       #STC_PH_xInitializeCard := TRUE;
       #STC_ST_xCardInitialized := FALSE;
   END_IF;
   #_w1 := #STC_ST_xRequestCardInitialization AND NOT #STC_ST_xPhaseInProgress AND NOT #STC_ST_xStoppingFaults AND NOT #INP_tHSCCount.ldStsSlot0;
   IF #_w1 THEN
       #STC_ST_xRequestCardInitialization := FALSE;
       #STC_AUX_tOutHSC.loadValue0 := 0;
   END_IF;
END_REGION

REGION Network 17: End initialize counter card
   RUNG wire#powerrail
      Contact( #STC_PH_xInitializeCard )
      wire#w1
      Contact( #STC_ST_xStoppingFaults )
      wire#w2
      R_Coil( #STC_PH_xInitializeCard )
   END_RUNG
   RUNG wire#w1
      Contact( #INP_tHSCCount.ldStsSlot0 )
   END_RUNG wire#w2
   RUNG wire#w2
      Coil( #STC_PH_xEndInitializeCard )
   END_RUNG
   // the same network as SCL:
   #_w1 := #STC_PH_xInitializeCard AND (#STC_ST_xStoppingFaults OR #INP_tHSCCount.ldStsSlot0);
   IF #_w1 THEN #STC_PH_xInitializeCard := FALSE; END_IF;
   #STC_PH_xEndInitializeCard := #_w1;
END_REGION

REGION Network 18: Set card initialized
   RUNG wire#powerrail
      Contact( #STC_PH_xEndInitializeCard )
      Contact( #INP_tHSCCount.ldStsSlot0 )
      I_Contact( #STC_ST_xStoppingFaults )
      wire#w1
      S_Coil( #STC_ST_xCardInitialized )
   END_RUNG
   RUNG wire#w1
      Coil( #TMP_xInitializeData )
   END_RUNG
   // the same network as SCL:
   #_w1 := #STC_PH_xEndInitializeCard AND #INP_tHSCCount.ldStsSlot0 AND NOT #STC_ST_xStoppingFaults;
   IF #_w1 THEN #STC_ST_xCardInitialized := TRUE; END_IF;
   #TMP_xInitializeData := #_w1;
END_REGION

REGION Network 19 (SCL): Initialize structure after initialization
   IF #TMP_xInitializeData THEN

       #INO_tEncoder.dActualEncoderCounter_cmm := 0;
       #INO_tEncoder.dLastMeterValue_cmm := 0;
       #INO_tEncoder.dNextMeterValue_cmm := #CONST_DMETERINC_CMM;
       #INO_tEncoder.rActSpeedValue_cmm_ms := 0.0;
       #STC_AUX_dLastCounterValue_cmm := 0;

       FOR #TMP_dIndex := 0 TO "DMAXXHEADS_IND" DO
           #INO_tEncoder.rgxMetersForXcuts[#TMP_dIndex] := FALSE;
       END_FOR;

       FOR #TMP_dIndex := 0 TO "DMAXYCUTBRIDGE_IND" DO
           #INO_tEncoder.rgxMetersForYCuts[#TMP_dIndex] := FALSE;
       END_FOR;

       #INO_tEncoder.xMeterForMarkers := FALSE;
       #INO_tEncoder.xMeterForScanner := FALSE;

       #STC_AUX_dLastMeterValue_cmm := 0;
       #STC_AUX_dNextMeterValue_cmm := #CONST_DMETERINC_CMM;
       #STC_AUX_lrTimingCounter_s := 0;
       #STC_AUX_lrTimingCounterFast_s := 0;
       #STC_AUX_dMeterValueSent_cmm := 0;

   END_IF;
END_REGION

REGION Network 20: ####_METER_THRESHOLD_####
END_REGION

REGION Network 21: Update new meter
   RUNG wire#powerrail
      Contact( #STC_ST_xCardInitialized )
      I_Contact( #STC_ST_xRequestCardInitialization )
      I_Contact( #STC_ST_xPhaseInProgress )
      I_Contact( #STC_ST_xStoppingFaults )
      I_Contact( #INP_tHSCCount.ldStsSlot0 )
      { S7_Templates := "SrcType := DInt" } NE_Contact(in1 := #STC_AUX_dNextMeterValue_cmm, in2 := #STC_AUX_dMeterValueSent_cmm)
      wire#w1
      S_Coil( #STC_PH_xUpdateNewMeter )
   END_RUNG
   RUNG wire#w1
      Move(in := #STC_AUX_dNextMeterValue_cmm, out1 => #STC_AUX_tOutHSC.loadValue0)
   END_RUNG
   // the same network as SCL:
   IF #STC_ST_xCardInitialized AND NOT #STC_ST_xRequestCardInitialization AND NOT #STC_ST_xPhaseInProgress AND NOT #STC_ST_xStoppingFaults AND NOT #INP_tHSCCount.ldStsSlot0 AND (#STC_AUX_dNextMeterValue_cmm <> #STC_AUX_dMeterValueSent_cmm) THEN
       #STC_PH_xUpdateNewMeter := TRUE;
       #STC_AUX_tOutHSC.loadValue0 := #STC_AUX_dNextMeterValue_cmm;
   END_IF;
END_REGION

REGION Network 22: End update new meter
   RUNG wire#powerrail
      Contact( #STC_PH_xUpdateNewMeter )
      wire#w1
      Contact( #INP_tHSCCount.ldStsSlot0 )
      wire#w2
      R_Coil( #STC_PH_xUpdateNewMeter )
   END_RUNG
   RUNG wire#w1
      Contact( #IN_xSimulationActive )
   END_RUNG wire#w2
   RUNG wire#w1
      Contact( #STC_ST_xStoppingFaults )
   END_RUNG wire#w2
   RUNG wire#w2
      Coil( #STC_PH_xEndUpdateNewMeter )
   END_RUNG
   // the same network as SCL:
   #_w1 := #STC_PH_xUpdateNewMeter AND (#INP_tHSCCount.ldStsSlot0 OR #IN_xSimulationActive OR #STC_ST_xStoppingFaults);
   IF #_w1 THEN #STC_PH_xUpdateNewMeter := FALSE; END_IF;
   #STC_PH_xEndUpdateNewMeter := #_w1;
END_REGION

REGION Network 23: Set meter correctly written
   RUNG wire#powerrail
      Contact( #STC_PH_xEndUpdateNewMeter )
      wire#w1
      Contact( #INP_tHSCCount.ldStsSlot0 )
      wire#w2
      Move(in := #STC_AUX_dNextMeterValue_cmm, out1 => #STC_AUX_dMeterValueSent_cmm)
   END_RUNG
   RUNG wire#w1
      Contact( #IN_xSimulationActive )
   END_RUNG wire#w2
   // the same network as SCL:
   IF #STC_PH_xEndUpdateNewMeter AND (#INP_tHSCCount.ldStsSlot0 OR #IN_xSimulationActive) THEN
       #STC_AUX_dMeterValueSent_cmm := #STC_AUX_dNextMeterValue_cmm;
   END_IF;
END_REGION

REGION Network 24: ####_NEW METER ARRIVED_####
END_REGION

REGION Network 25: Check if new meter arrived
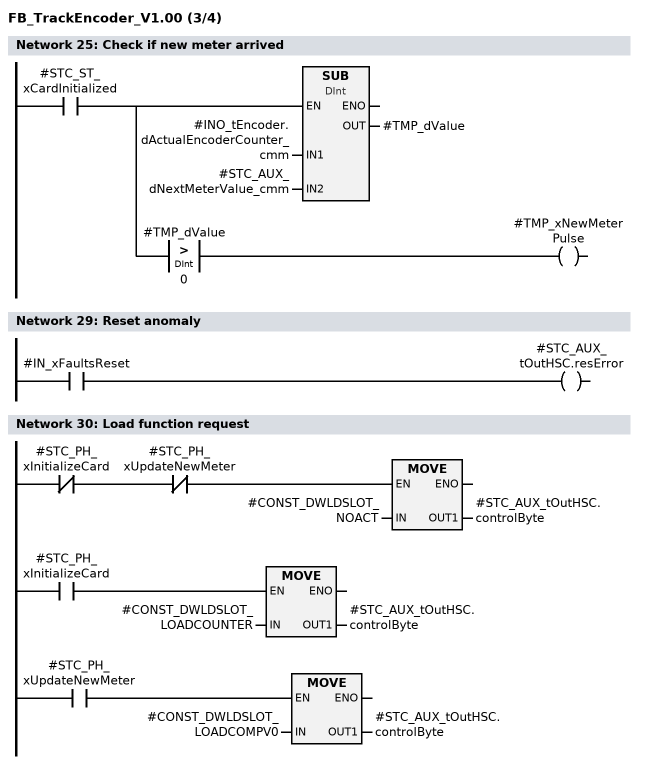
   RUNG wire#powerrail
      Contact( #STC_ST_xCardInitialized )
      wire#w1
      { S7_Templates := "SrcType := DInt" } Sub(in1 := #INO_tEncoder.dActualEncoderCounter_cmm, in2 := #STC_AUX_dNextMeterValue_cmm, out => #TMP_dValue)
   END_RUNG
   RUNG wire#w1
      { S7_Templates := "SrcType := DInt" } GT_Contact(in1 := #TMP_dValue, in2 := 0)
      Coil( #TMP_xNewMeterPulse )
   END_RUNG
   // the same network as SCL:
   IF #STC_ST_xCardInitialized THEN
       #TMP_dValue := #INO_tEncoder.dActualEncoderCounter_cmm - #STC_AUX_dNextMeterValue_cmm;
   END_IF;
   #TMP_xNewMeterPulse := #STC_ST_xCardInitialized AND (#TMP_dValue > 0);
END_REGION

REGION Network 26 (SCL): New meter pulse
   IF #TMP_xNewMeterPulse THEN

       #STC_AUX_dLastMeterValue_cmm := #STC_AUX_dNextMeterValue_cmm;
       #STC_AUX_dNextMeterValue_cmm += #CONST_DMETERINC_CMM;

       #INO_tEncoder.dLastMeterValue_cmm := #STC_AUX_dLastMeterValue_cmm; 
       #INO_tEncoder.dNextMeterValue_cmm := #STC_AUX_dNextMeterValue_cmm; 

       FOR #TMP_dIndex := 0 TO "DMAXXHEADS_IND" DO
           #INO_tEncoder.rgxMetersForXcuts[#TMP_dIndex] := TRUE;
       END_FOR;

       FOR #TMP_dIndex := 0 TO "DMAXYCUTBRIDGE_IND" DO
           #INO_tEncoder.rgxMetersForYCuts[#TMP_dIndex] := TRUE;
       END_FOR;

       #INO_tEncoder.xMeterForMarkers := TRUE;
       #INO_tEncoder.xMeterForScanner := TRUE;


   END_IF;
END_REGION

REGION Network 27 (SCL): Calculate speed
   #STC_AUX_lrTimingCounter_s += #STC_AUX_lrElapsedTime_s;
   #STC_AUX_lrTimingCounterFast_s += #STC_AUX_lrElapsedTime_s;

   IF #STC_AUX_lrTimingCounter_s >= #CONST_LRUPDATESPEED_S THEN

       #TMP_dElapsedPulses_cmm := #INO_tEncoder.dActualEncoderCounter_cmm - #STC_AUX_dLastCounterValue_cmm;

       #INO_tEncoder.rActSpeedValue_cmm_ms := DINT_TO_REAL(#TMP_dElapsedPulses_cmm) / (LREAL_TO_REAL(#STC_AUX_lrTimingCounter_s) * 1000.0);
       #INO_tEncoder.dActSpeedValue_mm_min := REAL_TO_DINT(#INO_tEncoder.rActSpeedValue_cmm_ms * 600.0);    

       #STC_AUX_dLastCounterValue_cmm := #INO_tEncoder.dActualEncoderCounter_cmm;
       #STC_AUX_lrTimingCounter_s := 0;

   END_IF;

   IF #STC_AUX_lrTimingCounterFast_s >= #CONST_LRUPDATESPEEDFAST_S THEN

       #TMP_dElapsedPulses_cmm := #INO_tEncoder.dActualEncoderCounter_cmm - #STC_AUX_dLastCounterValueFast_cmm;

       #INO_tEncoder.rActSpeedValueFast_cmm_ms := DINT_TO_REAL(#TMP_dElapsedPulses_cmm) / (LREAL_TO_REAL(#STC_AUX_lrTimingCounterFast_s) * 1000.0);
       #INO_tEncoder.dActSpeedValueFast_mm_min := REAL_TO_DINT(#INO_tEncoder.rActSpeedValueFast_cmm_ms * 600.0);    

       #STC_AUX_dLastCounterValueFast_cmm := #INO_tEncoder.dActualEncoderCounter_cmm;
       #STC_AUX_lrTimingCounterFast_s := 0;

   END_IF;
END_REGION

REGION Network 28: ####_OUTPUT_####
END_REGION

REGION Network 29: Reset anomaly
   RUNG wire#powerrail
      Contact( #IN_xFaultsReset )
      Coil( #STC_AUX_tOutHSC.resError )
   END_RUNG
   // the same network as SCL:
   #STC_AUX_tOutHSC.resError := #IN_xFaultsReset;
END_REGION

REGION Network 30: Load function request
   RUNG wire#powerrail
      I_Contact( #STC_PH_xInitializeCard )
      I_Contact( #STC_PH_xUpdateNewMeter )
      Move(in := #CONST_DWLDSLOT_NOACT, out1 => #STC_AUX_tOutHSC.controlByte)
   END_RUNG
   RUNG wire#powerrail
      Contact( #STC_PH_xInitializeCard )
      Move(in := #CONST_DWLDSLOT_LOADCOUNTER, out1 => #STC_AUX_tOutHSC.controlByte)
   END_RUNG
   RUNG wire#powerrail
      Contact( #STC_PH_xUpdateNewMeter )
      Move(in := #CONST_DWLDSLOT_LOADCOMPV0, out1 => #STC_AUX_tOutHSC.controlByte)
   END_RUNG
   // the same network as SCL:
   IF NOT #STC_PH_xInitializeCard AND NOT #STC_PH_xUpdateNewMeter THEN
       #STC_AUX_tOutHSC.controlByte := #CONST_DWLDSLOT_NOACT;
   END_IF;
   IF #STC_PH_xInitializeCard THEN #STC_AUX_tOutHSC.controlByte := #CONST_DWLDSLOT_LOADCOUNTER; END_IF;
   IF #STC_PH_xUpdateNewMeter THEN #STC_AUX_tOutHSC.controlByte := #CONST_DWLDSLOT_LOADCOMPV0; END_IF;
END_REGION

REGION Network 31: Fixed command
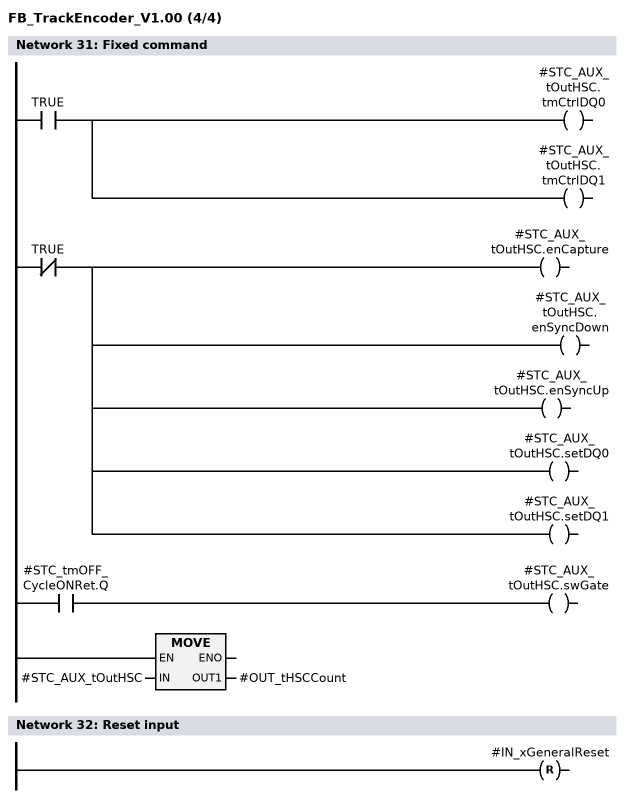
   RUNG wire#powerrail
      Contact( TRUE )
      wire#w1
      Coil( #STC_AUX_tOutHSC.tmCtrlDQ0 )
   END_RUNG
   RUNG wire#w1
      Coil( #STC_AUX_tOutHSC.tmCtrlDQ1 )
   END_RUNG
   RUNG wire#powerrail
      I_Contact( TRUE )
      wire#w2
      Coil( #STC_AUX_tOutHSC.enCapture )
   END_RUNG
   RUNG wire#w2
      Coil( #STC_AUX_tOutHSC.enSyncDown )
   END_RUNG
   RUNG wire#w2
      Coil( #STC_AUX_tOutHSC.enSyncUp )
   END_RUNG
   RUNG wire#w2
      Coil( #STC_AUX_tOutHSC.setDQ0 )
   END_RUNG
   RUNG wire#w2
      Coil( #STC_AUX_tOutHSC.setDQ1 )
   END_RUNG
   RUNG wire#powerrail
      Contact( #STC_tmOFF_CycleONRet.Q )
      Coil( #STC_AUX_tOutHSC.swGate )
   END_RUNG
   RUNG wire#powerrail
      Move(in := #STC_AUX_tOutHSC, out1 => #OUT_tHSCCount)
   END_RUNG
   // the same network as SCL:
   #STC_AUX_tOutHSC.tmCtrlDQ0 := TRUE;
   #STC_AUX_tOutHSC.tmCtrlDQ1 := TRUE;
   #STC_AUX_tOutHSC.enCapture := NOT TRUE;
   #STC_AUX_tOutHSC.enSyncDown := NOT TRUE;
   #STC_AUX_tOutHSC.enSyncUp := NOT TRUE;
   #STC_AUX_tOutHSC.setDQ0 := NOT TRUE;
   #STC_AUX_tOutHSC.setDQ1 := NOT TRUE;
   #STC_AUX_tOutHSC.swGate := #STC_tmOFF_CycleONRet.Q;
   #OUT_tHSCCount := #STC_AUX_tOutHSC;
END_REGION

REGION Network 32: Reset input
   RUNG wire#powerrail
      R_Coil( #IN_xGeneralReset )
   END_RUNG
   // the same network as SCL:
   #IN_xGeneralReset := FALSE;
END_REGION
END_FUNCTION_BLOCK

// folder: 03_Programs_Logics/MCC1200/05_ExternalOPT

FUNCTION_BLOCK "FB_OptManager_V1.00"   // FB6, LAD
{ S7_Optimized_Access := 'TRUE' }
VERSION : 0.1
   VAR_INPUT
      IN_xFaultsEnabled : Bool;   // Faults enabled
      IN_xCycleON : Bool;   // Zone is in cycle
      IN_xGeneralReset : Bool;   // General reset
      IN_xFaultsReset : Bool;   // Reset alarms
      IN_dGlassDataMachineIndex : DInt;   // Glass data machine index
      IN_dGlassDataRequestMachineIndex : DInt;   // Glass data request machine index
      IN_dGlassDataUpdateMachineIndex : DInt;   // Glass data update machine index
   END_VAR
   VAR_IN_OUT
      INO_tCaps : "UDT_CapData_Tracking";   // Cap tracking
      INO_tEncoder : "UDT_Encoder";   // Encoder data
      INO_tRibbon : "UDT_RibbonData";   // Ribbon data
      INO_tDefects : "UDT_DefectData_Tracking_Ext";   // Defects data
   END_VAR
   VAR RETAIN
      tHMW : Struct   // HMI Write
         dDecisionLinePosition_cmm : DInt;   // Decision line position [mm/100] {mm/100|mm|0|30000|M}
         dLastOptLinePosition_cmm : DInt;   // Last optimizer line position [mm/100] {mm/100|mm|0|30000|M}
         dSelectRibbonDataSource : DInt;   // Select ribbon data source (0=Manual 1=Scanner 2=Camera) {X|X|0|2|O}
         dSelectWanderDataSource : DInt;   // Select wander data source (0=Manual 1=Scanner 2=Camera) {X|X|0|2|O}
         dSelectWanderMode : DInt;   // Select wander mode (0=Net 1=Gross)
         dManualGrossWidth_cmm : DInt;   // Manual gross width [mm/100] {mm/100|mm|2000|4000|O}
         dManualNetWidth_cmm : DInt;   // Manual net width [mm/100] {mm/100|mm|2000|4000|O}
         dManualWander_cmm : DInt;   // Manual wander [mm/100] {mm/100|mm|-200|200|O}
         dWanderOffset_cmm : DInt;   // Wander offset [mm/100] {mm/100|mm|-200|200|O}
         dWanderRecThr_cmm : DInt;   // Wander recovery threshold [mm/100] {mm/100|mm|-200|200|O}
         xUpdateLastOptimizerLine : Bool;   // Update last optimizer line position {X|X|X|X|M}
         xUpdateDecisionLine : Bool;   // Update decision line position {X|X|X|X|M}
         xSelectOptimizerA : Bool;   // Select optimizer A {X|X|X|X|O}
         xSelectOptimizerB : Bool;   // Select optimizer B {X|X|X|X|O}
      END_STRUCT;
      tHMR : Struct   // HMI Read
         dLastOptLinePosition_cmm : DInt;   // Last optimizer line position [mm/100]
         dDecisionLinePosition_cmm : DInt;   // Decision line position [mm/100]
         dSelOptimizer : DInt;   // Selected optimizer (1= OptA 2=OptB)
         rgtRibbonData : Array[0.."DMAXGLASSDATAMACHINE_IND"] of Struct
            dGrossWidth_cmm : DInt;   // Gross width [mm/100]
            dNetWidth_cmm : DInt;   // Net width [mm/100]
            dGrossWander_cmm : DInt;   // Gross wander [mm/100]
            dNetWander_cmm : DInt;   // Net wander [mm/100]
         END_STRUCT;
      END_STRUCT;
   END_VAR
   VAR
      OSR_xGeneralReset : Bool;   // General reset
      AUX_dLastGlassDataUpdated : DInt;   // Last index glass data update
   END_VAR
   VAR_TEMP
      TMP_xOSGeneralReset : Bool;
      TMP_dIndex : DInt;
      TMP_dID : DInt;
      TMP_xManualDataIsChanged : Bool;   // Manual data is changed
      TMP_dwMask : DWord;
      TMP_wMask : Word;
      AUX_dNumPlatePacket : DInt;
      TMP_iReturn : Int;
      TMP_dTargetTest : DInt;
      TMP_xRandOut : Bool;
      TMP_wStatus : Word;
      TMP_dLength : DInt;
   END_VAR
   VAR_TEMP   // added for the SCL form of the ladder/FBD networks
      _w1 : Bool;
   END_VAR
BEGIN

REGION Network 3: Calculate OS of the general reset
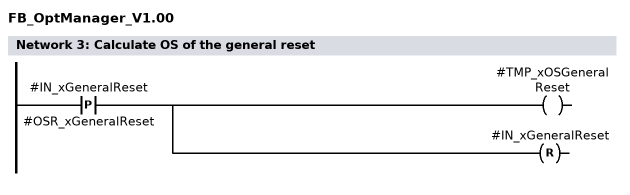
   RUNG wire#powerrail
      P_Contact(operand := #IN_xGeneralReset, bit := #OSR_xGeneralReset)
      wire#w1
      Coil( #TMP_xOSGeneralReset )
   END_RUNG
   RUNG wire#w1
      R_Coil( #IN_xGeneralReset )
   END_RUNG
   // the same network as SCL:
   #_w1 := #IN_xGeneralReset AND NOT #OSR_xGeneralReset;   // rising edge of #IN_xGeneralReset
   #OSR_xGeneralReset := #IN_xGeneralReset;
   #TMP_xOSGeneralReset := #_w1;
   IF #_w1 THEN #IN_xGeneralReset := FALSE; END_IF;
END_REGION

REGION Network 4 (SCL): General reset
   #INO_tCaps.rgtTrackMachine["DMACHINEINDEX_LASTOPTLINE"].tUserData.dSetDistanceSnap_cmm := #tHMR.dLastOptLinePosition_cmm;
   #INO_tCaps.rgtTrackMachine["DMACHINEINDEX_LASTOPTLINE"].tUserData.dSetMachReacTime_ms := 0;

   IF #TMP_xOSGeneralReset THEN

       #INO_tCaps.rgtTrackMachine["DMACHINEINDEX_LASTOPTLINE"].tUserData.dSetDistanceSnap_cmm := #tHMR.dLastOptLinePosition_cmm;
       #INO_tCaps.rgtTrackMachine["DMACHINEINDEX_LASTOPTLINE"].tUserData.dSetMachReacTime_ms := 0;
       #INO_tRibbon.rgtGlassData[#IN_dGlassDataMachineIndex].dDistSnapRoll_cmm := #tHMR.dDecisionLinePosition_cmm;

       #AUX_dLastGlassDataUpdated := 0;

       #INO_tRibbon.rgtGlassDataUpdate[#IN_dGlassDataUpdateMachineIndex].tData.dGrossWidth_cmm := 0;
       #INO_tRibbon.rgtGlassDataUpdate[#IN_dGlassDataUpdateMachineIndex].tData.dNetWidth_cmm := 0;
       #INO_tRibbon.rgtGlassDataUpdate[#IN_dGlassDataUpdateMachineIndex].tData.dGrossWander_cmm := 0;
       #INO_tRibbon.rgtGlassDataUpdate[#IN_dGlassDataUpdateMachineIndex].tData.dNetWander_cmm := 0;

   END_IF;
END_REGION

REGION Network 5 (SCL): #### HMI LOGICS ####
   IF #tHMW.xUpdateLastOptimizerLine THEN
       #tHMW.xUpdateLastOptimizerLine := FALSE;
       #tHMR.dLastOptLinePosition_cmm := #tHMW.dLastOptLinePosition_cmm;
       #INO_tCaps.rgtTrackMachine["DMACHINEINDEX_LASTOPTLINE"].tUserData.dSetDistanceSnap_cmm := #tHMR.dLastOptLinePosition_cmm;
   END_IF;

   IF #tHMW.xUpdateDecisionLine THEN
       #tHMW.xUpdateDecisionLine := FALSE;
       #tHMR.dDecisionLinePosition_cmm := #tHMW.dDecisionLinePosition_cmm;
       #INO_tRibbon.rgtGlassData[#IN_dGlassDataMachineIndex].dDistSnapRoll_cmm := #tHMR.dDecisionLinePosition_cmm;
   END_IF;

   IF #INO_tRibbon.rgtGlassDataRequest[#IN_dGlassDataRequestMachineIndex].OUT_xDataReady THEN

       #tHMR.rgtRibbonData[#AUX_dLastGlassDataUpdated].dGrossWander_cmm := #INO_tRibbon.rgtGlassDataRequest[#IN_dGlassDataRequestMachineIndex].OUT_dGrossWander_cmm;
       #tHMR.rgtRibbonData[#AUX_dLastGlassDataUpdated].dGrossWidth_cmm := #INO_tRibbon.rgtGlassDataRequest[#IN_dGlassDataRequestMachineIndex].OUT_dGrossWidth_cmm;
       #tHMR.rgtRibbonData[#AUX_dLastGlassDataUpdated].dNetWander_cmm := #INO_tRibbon.rgtGlassDataRequest[#IN_dGlassDataRequestMachineIndex].OUT_dNetWander_cmm;
       #tHMR.rgtRibbonData[#AUX_dLastGlassDataUpdated].dNetWidth_cmm := #INO_tRibbon.rgtGlassDataRequest[#IN_dGlassDataRequestMachineIndex].OUT_dNetWidth_cmm;

   END_IF;

   //Retrieve the value of ribbon near the decision line position
   IF NOT #INO_tRibbon.rgtGlassDataRequest[#IN_dGlassDataRequestMachineIndex].IN_xRequestGlassData OR #INO_tRibbon.rgtGlassDataRequest[#IN_dGlassDataRequestMachineIndex].OUT_xDataReady THEN

       #INO_tRibbon.rgtGlassDataRequest[#IN_dGlassDataRequestMachineIndex].OUT_xDataReady := FALSE;

       #AUX_dLastGlassDataUpdated += 1;

       IF (#AUX_dLastGlassDataUpdated > #INO_tRibbon.dActualNumberGlassDataMachine - 1) THEN
           #AUX_dLastGlassDataUpdated := 0;
       END_IF;

       #INO_tRibbon.rgtGlassDataRequest[#IN_dGlassDataRequestMachineIndex].IN_dDistanceSnaproll_cmm := #tHMR.dDecisionLinePosition_cmm;
       #INO_tRibbon.rgtGlassDataRequest[#IN_dGlassDataRequestMachineIndex].IN_dSourceIndex := #AUX_dLastGlassDataUpdated;
       #INO_tRibbon.rgtGlassDataRequest[#IN_dGlassDataRequestMachineIndex].IN_xRequestGlassData := TRUE;

   END_IF;

   //Update the manual glass data selection 
   IF #tHMW.dSelectRibbonDataSource > 0 THEN
       #tHMW.dManualGrossWidth_cmm := #tHMR.rgtRibbonData[#tHMW.dSelectRibbonDataSource].dGrossWidth_cmm;
       #tHMW.dManualNetWidth_cmm := #tHMR.rgtRibbonData[#tHMW.dSelectRibbonDataSource].dNetWidth_cmm;
   END_IF;

   //Update the manual glass data selection
   IF #tHMW.dSelectWanderDataSource > 0 THEN
       #tHMW.dManualWander_cmm := #tHMR.rgtRibbonData[#tHMW.dSelectWanderDataSource].dNetWander_cmm;
   END_IF;

   #TMP_xManualDataIsChanged := FALSE;

   //Check if some data are changed
   IF ((#tHMW.dManualWander_cmm <> #INO_tRibbon.rgtGlassDataUpdate[#IN_dGlassDataUpdateMachineIndex].tData.dGrossWander_cmm) OR
       (#tHMW.dManualWander_cmm <> #INO_tRibbon.rgtGlassDataUpdate[#IN_dGlassDataUpdateMachineIndex].tData.dNetWander_cmm) OR
       (#tHMW.dManualGrossWidth_cmm <> #INO_tRibbon.rgtGlassDataUpdate[#IN_dGlassDataUpdateMachineIndex].tData.dGrossWidth_cmm) OR
       (#tHMW.dManualNetWidth_cmm <> #INO_tRibbon.rgtGlassDataUpdate[#IN_dGlassDataUpdateMachineIndex].tData.dNetWidth_cmm)) THEN

       #TMP_xManualDataIsChanged := TRUE;

   END_IF;

   //Update the manual data buffer
   IF NOT #INO_tRibbon.rgtGlassDataUpdate[#IN_dGlassDataUpdateMachineIndex].xUpdateRequest AND #TMP_xManualDataIsChanged  THEN
       #INO_tRibbon.rgtGlassDataUpdate[#IN_dGlassDataUpdateMachineIndex].tData.dGrossWander_cmm := #tHMW.dManualWander_cmm;
       #INO_tRibbon.rgtGlassDataUpdate[#IN_dGlassDataUpdateMachineIndex].tData.dNetWander_cmm := #tHMW.dManualWander_cmm;
       #INO_tRibbon.rgtGlassDataUpdate[#IN_dGlassDataUpdateMachineIndex].tData.dGrossWidth_cmm := #tHMW.dManualGrossWidth_cmm;
       #INO_tRibbon.rgtGlassDataUpdate[#IN_dGlassDataUpdateMachineIndex].tData.dNetWidth_cmm := #tHMW.dManualNetWidth_cmm;

       #INO_tRibbon.rgtGlassDataUpdate[#IN_dGlassDataUpdateMachineIndex].xUpdateRequest := TRUE;

   END_IF;

   IF #tHMW.xSelectOptimizerA THEN
       #tHMR.dSelOptimizer := 1;
       #tHMW.xSelectOptimizerA := FALSE;
   END_IF;

   IF #tHMW.xSelectOptimizerB THEN
       #tHMR.dSelOptimizer := 2;
       #tHMW.xSelectOptimizerB := FALSE;
   END_IF;
END_REGION

REGION Network 6 (SCL): Insert plate in case of timeout plate on tracking buffer
   //Update the data of the last target line
   #INO_tCaps.rgtTrackMachine["DMACHINEINDEX_LASTOPTLINE"].tUserData.dSetMachReacTime_ms := 0;

   #TMP_dTargetTest := #INO_tCaps.dLastTargetLineValue_cmm - #INO_tEncoder.dActualEncoderCounter_cmm; 

   IF #INO_tCaps.rgtTrackMachine["DMACHINEINDEX_LASTOPTLINE"].tUserData.xGetPosReach
   (* OR 
       ("GP_OB_Initialize_Medium_IDB".OUT_xOs_30s AND #TMP_dTargetTest > 100000 AND #INO_tEncoder.dActSpeedValue_mm_min > 1000)*)  THEN

       #TMP_dLength :=  "LGF_RandomRange_Dint"(minValue:=15000, maxValue:=30000, error=>#TMP_xRandOut, subfunctionStatus=>#TMP_wStatus, status=>#TMP_wStatus);

       #INO_tCaps.tNewCapToInsert.dID := #INO_tCaps.dNextValidCapID;
       #TMP_dID := #INO_tCaps.dNextValidCapID + 1;
       IF #INO_tCaps.rgtTrackMachine["DMACHINEINDEX_LASTOPTLINE"].tUserData.xGetPosReach THEN
           #INO_tCaps.tNewCapToInsert.dLength_cmm := 200000;
       ELSE
           #INO_tCaps.tNewCapToInsert.dLength_cmm := #TMP_dLength;
       END_IF;

       FOR #TMP_dIndex := 0 TO #INO_tCaps.tNewCapToInsert.dNumLites - 1 DO
           #INO_tCaps.tNewCapToInsert.rgtLites[#TMP_dIndex].dMainDestination := "DCULLETDESTMASK";

           #INO_tCaps.tNewCapToInsert.rgtLites[#TMP_dIndex].dAltDestination := 0;
           #INO_tCaps.tNewCapToInsert.rgtLites[#TMP_dIndex].d2ndDestionation := 0;

           #INO_tCaps.tNewCapToInsert.rgtLites[#TMP_dIndex].dCulletCause := "DCULLETCAUSE_CAPDATATIMEOUT";
           #INO_tCaps.tNewCapToInsert.rgtLites[#TMP_dIndex].dProductionID := 0;
           #INO_tCaps.tNewCapToInsert.rgtLites[#TMP_dIndex].dID := #TMP_dID;

           #TMP_dID += 1;                        
       END_FOR;

       #INO_tCaps.tNewCapToInsert.tRequests.rgxXCutReqHead[0]:= TRUE;
       #INO_tCaps.tNewCapToInsert.tRequests.rgxXCutReqHead[1]:= TRUE;
       #INO_tCaps.tNewCapToInsert.tRequests.rgxXCutReqHead[2]:= TRUE;
       #INO_tCaps.tNewCapToInsert.tRequests.rgxXCutReqHead[3]:= TRUE;

       #INO_tCaps.tNewCapToInsert.tRequests.rgxXCutReqTail[0]:= TRUE;
       #INO_tCaps.tNewCapToInsert.tRequests.rgxXCutReqTail[1]:= TRUE;
       #INO_tCaps.tNewCapToInsert.tRequests.rgxXCutReqTail[2]:= TRUE;
       #INO_tCaps.tNewCapToInsert.tRequests.rgxXCutReqTail[3]:= TRUE;

       #INO_tCaps.tNewCapToInsert.tRequests.tYCutsData[0].xUseThisBridge:= FALSE;
       #INO_tCaps.tNewCapToInsert.tRequests.tYCutsData[1].xUseThisBridge:= FALSE;

       #INO_tCaps.tNewCapToInsert.tRequests.xUpdateDataBPSA := TRUE;    
       #INO_tCaps.tNewCapToInsert.tRequests.xUpdateDataBPSB := TRUE;    

       #INO_tCaps.xInsertCapOnTrack := TRUE;
       #INO_tCaps.rgtTrackMachine["DMACHINEINDEX_LASTOPTLINE"].tUserData.xGetPosReach := FALSE;

   END_IF;
END_REGION

REGION Network 7 (SCL): Manage internal PLC optimizer
   //Update the data for the optimizer
   (*"DB_OPTPLC_ExchangeData".TrackingData.dActualEncoderCounter_cmm := #INO_tEncoder.dActualEncoderCounter_cmm;
   "DB_OPTPLC_ExchangeData".TrackingData.dLastPlateID := #INO_tCaps.dLastValidCapID;
   "DB_OPTPLC_ExchangeData".TrackingData.dLastTargetLine_cmm := #INO_tCaps.dLastTargetLineValue_cmm;
   "DB_OPTPLC_ExchangeData".TrackingData.dOptDecisionLine_cmm := #tHMR.dDecisionLinePosition_cmm;

   //Evaluate the PLC optimizer response. In case of data valid, place the data inside the buffer
   IF "DB_OPTPLC_ExchangeData".PlcOptData.xCapDataReady 
       AND TRUE 
       AND "DB_OPTPLC_ExchangeData".PlcOptData.AUX_tPlatePacket.dPlateHead_cmm = #INO_tCaps.dLastTargetLineValue_cmm
       AND "DB_OPTPLC_ExchangeData".PlcOptData.AUX_tPlatePacket.dCapID = #INO_tCaps.dNextValidCapID THEN

       #INO_tCaps.tNewCapToInsert := #INO_tCaps.tEmptyCap;

       #INO_tCaps.tNewCapToInsert.dID := "DB_OPTPLC_ExchangeData".PlcOptData.AUX_tPlatePacket.dCapID;
       #INO_tCaps.tNewCapToInsert.dHeadPositionBTC := "DB_OPTPLC_ExchangeData".PlcOptData.AUX_tPlatePacket.dPlateHead_cmm;
       #INO_tCaps.tNewCapToInsert.dTailPositionBTC := #INO_tCaps.tNewCapToInsert.dHeadPositionBTC + "DB_OPTPLC_ExchangeData".PlcOptData.AUX_tPlatePacket.dCapLength_cmm;
       #INO_tCaps.tNewCapToInsert.dLength_cmm := "DB_OPTPLC_ExchangeData".PlcOptData.AUX_tPlatePacket.dCapLength_cmm;
       #INO_tCaps.tNewCapToInsert.dWidth_cmm := "DB_OPTPLC_ExchangeData".PlcOptData.AUX_tPlatePacket.dTotCapWidth_cmm;
       #INO_tCaps.tNewCapToInsert.dThick_cmm := "DB_OPTPLC_ExchangeData".PlcOptData.AUX_tPlatePacket.dCapThick_cmm;
       #INO_tCaps.tNewCapToInsert.dIndex := "DB_OPTPLC_ExchangeData".PlcOptData.AUX_tPlatePacket.dIndexPlateConv;
       #INO_tCaps.tNewCapToInsert.dFormat := 0;
       #INO_tCaps.tNewCapToInsert.dNumLites := "DB_OPTPLC_ExchangeData".PlcOptData.AUX_tPlatePacket.dNumLiteCap;
       #INO_tCaps.tNewCapToInsert.dReqGapForConv_cmm := 0;
       #INO_tCaps.tNewCapToInsert.dMaxCapInConv := "DB_OPTPLC_ExchangeData".PlcOptData.AUX_tPlatePacket.dMaxPlateConv;
       #INO_tCaps.tNewCapToInsert.dConvTotLength_cmm := "DB_OPTPLC_ExchangeData".PlcOptData.AUX_tPlatePacket.dConvLength_cmm;
       #INO_tCaps.tNewCapToInsert.dMinWidth_cmm := "DB_OPTPLC_ExchangeData".PlcOptData.AUX_tPlatePacket.dMinWidth_cmm;
       #INO_tCaps.tNewCapToInsert.dMaxWidth_cmm := "DB_OPTPLC_ExchangeData".PlcOptData.AUX_tPlatePacket.dMaxWidth_cmm;
       #INO_tCaps.tNewCapToInsert.dGrossWidth_cmm := 0;
       #INO_tCaps.tNewCapToInsert.dNetWidth_cmm := 0;
       #INO_tCaps.tNewCapToInsert.dDEdgeOpSide_cmm := "DB_OPTPLC_ExchangeData".PlcOptData.AUX_tPlatePacket.dExtBordOp;
       #INO_tCaps.tNewCapToInsert.dDEdgeOppOpSide_cmm := "DB_OPTPLC_ExchangeData".PlcOptData.AUX_tPlatePacket.dExtBordOppoOp;
       #INO_tCaps.tNewCapToInsert.dTEdgeOpSide_cmm := 0;
       #INO_tCaps.tNewCapToInsert.dTEdgeOppOpSide_cmm := 0;
       #INO_tCaps.tNewCapToInsert.dStartCutWander_cmm := "DB_OPTPLC_ExchangeData".PlcOptData.AUX_tPlatePacket.dWanderRec_cmm;
       #INO_tCaps.tNewCapToInsert.dEndCutWander_cmm := "DB_OPTPLC_ExchangeData".PlcOptData.AUX_tPlatePacket.dWanderRec_cmm;
       #INO_tCaps.tNewCapToInsert.dNetWander_cmm := 0;
       #INO_tCaps.tNewCapToInsert.dGrossWander_cmm := 0;
       #INO_tCaps.tNewCapToInsert.dColor := "DB_OPTPLC_ExchangeData".PlcOptData.AUX_tPlatePacket.dColorID;
       #INO_tCaps.tNewCapToInsert.strColorDescr := '';
       #INO_tCaps.tNewCapToInsert.dSystemMeasure := 0;

       IF "DB_OPTPLC_ExchangeData".PlcOptData.AUX_tPlatePacket.dYBridgeToCut = 1 THEN

           #INO_tCaps.tNewCapToInsert.tRequests.tYCutsData[0].rgdHeadsPositions := "DB_OPTPLC_ExchangeData".PlcOptData.AUX_tPlatePacket.rgYBridgePos_cmm;

           GATHER(IN:="DB_OPTPLC_ExchangeData".PlcOptData.AUX_tPlatePacket.rgxYHeadMask,
                  OUT=>#TMP_dwMask);

           #TMP_wMask := DWORD_TO_WORD(#TMP_dwMask);     

           SCATTER(IN:=#TMP_wMask,
                   OUT=>#INO_tCaps.tNewCapToInsert.tRequests.tYCutsData[0].rgxHeadsRequest);

           #INO_tCaps.tNewCapToInsert.tRequests.tYCutsData[0].xUseThisBridge := TRUE;

       ELSIF "DB_OPTPLC_ExchangeData".PlcOptData.AUX_tPlatePacket.dYBridgeToCut = 2 THEN

           #INO_tCaps.tNewCapToInsert.tRequests.tYCutsData[1].rgdHeadsPositions := "DB_OPTPLC_ExchangeData".PlcOptData.AUX_tPlatePacket.rgYBridgePos_cmm;

           GATHER(IN:="DB_OPTPLC_ExchangeData".PlcOptData.AUX_tPlatePacket.rgxYHeadMask,
                  OUT=>#TMP_dwMask);

           #TMP_wMask := DWORD_TO_WORD(#TMP_dwMask);     

           SCATTER(IN:=#TMP_wMask,
                   OUT=>#INO_tCaps.tNewCapToInsert.tRequests.tYCutsData[1].rgxHeadsRequest);

           #INO_tCaps.tNewCapToInsert.tRequests.tYCutsData[1].xUseThisBridge := TRUE;

       END_IF;

       FOR #TMP_dIndex := 0 TO "DMAXXHEADS_IND" DO

           #INO_tCaps.tNewCapToInsert.tRequests.rgxXCutReqHead[#TMP_dIndex] := TRUE;//#AUX_rgtPlatePacketArray[0].rgxCutMissionHead[#TMP_dIndex];
           #INO_tCaps.tNewCapToInsert.tRequests.rgxXCutReqTail[#TMP_dIndex] := TRUE;//#AUX_rgtPlatePacketArray[0].rgxCutMissionTail[#TMP_dIndex];

       END_FOR;

       #INO_tCaps.tNewCapToInsert.tRequests.xOptSelvedgeSel := NOT "DB_OPTPLC_ExchangeData".PlcOptData.AUX_tPlatePacket.tGeneralFlags.xAutoTrim;
       #INO_tCaps.tNewCapToInsert.tRequests.xOptSplitBarSel := NOT "DB_OPTPLC_ExchangeData".PlcOptData.AUX_tPlatePacket.tGeneralFlags.xAutoSnap;
       #INO_tCaps.tNewCapToInsert.tRequests.xOptSepRollSel := NOT "DB_OPTPLC_ExchangeData".PlcOptData.AUX_tPlatePacket.tGeneralFlags.xAutoSep;
       #INO_tCaps.tNewCapToInsert.tRequests.dReqTrim3OpSide := 0;
       #INO_tCaps.tNewCapToInsert.tRequests.dReqTrim2OpSide := "DB_OPTPLC_ExchangeData".PlcOptData.AUX_tPlatePacket.dExtBordOp;
       #INO_tCaps.tNewCapToInsert.tRequests.dReqTrim1OpSide :=  "DB_OPTPLC_ExchangeData".PlcOptData.AUX_tPlatePacket.dIntBordOp;
       #INO_tCaps.tNewCapToInsert.tRequests.dReqTrim3OppOpSide := 0;
       #INO_tCaps.tNewCapToInsert.tRequests.dReqTrim2OppOpSide := "DB_OPTPLC_ExchangeData".PlcOptData.AUX_tPlatePacket.dExtBordOppoOp;
       #INO_tCaps.tNewCapToInsert.tRequests.dReqTrim1OppOpSide := "DB_OPTPLC_ExchangeData".PlcOptData.AUX_tPlatePacket.dIntBordOp;
       #INO_tCaps.tNewCapToInsert.tRequests.rgdReqSplitBarSel := "DB_OPTPLC_ExchangeData".PlcOptData.AUX_tPlatePacket.rgdBumps;

       GATHER(IN:="DB_OPTPLC_ExchangeData".PlcOptData.AUX_tPlatePacket.rgxChevrons,
              OUT=>#TMP_dwMask);

       #INO_tCaps.tNewCapToInsert.tRequests.rgbSeparatorSelect[0] := DWORD_TO_BYTE(SHR(IN:=#TMP_dwMask, N:=24));
       #INO_tCaps.tNewCapToInsert.tRequests.rgbSeparatorSelect[1] := DWORD_TO_BYTE(SHR(IN:=SHL(IN:=#TMP_dwMask,N:= 8), N:=24));
       #INO_tCaps.tNewCapToInsert.tRequests.rgbSeparatorSelect[2] := DWORD_TO_BYTE(SHR(IN:=SHL(IN:=#TMP_dwMask,N:= 16), N:=24));
       #INO_tCaps.tNewCapToInsert.tRequests.rgbSeparatorSelect[3] := DWORD_TO_BYTE(SHR(IN:=SHL(IN:=#TMP_dwMask,N:= 24), N:=24));

       #INO_tCaps.tNewCapToInsert.tRequests.xUpdateDataBPSA := TRUE;
       #INO_tCaps.tNewCapToInsert.tRequests.xUpdateDataBPSB := TRUE;
       #INO_tCaps.tNewCapToInsert.tRequests.xWandContinue := TRUE;

       FOR #TMP_dIndex := 0 TO "DB_OPTPLC_ExchangeData".PlcOptData.AUX_tPlatePacket.dNumLiteCap - 1 DO

           #INO_tCaps.tNewCapToInsert.rgtLites[#TMP_dIndex].dID := "DB_OPTPLC_ExchangeData".PlcOptData.AUX_tPlatePacket.rgdLiteID[#TMP_dIndex];
           #INO_tCaps.tNewCapToInsert.rgtLites[#TMP_dIndex].dProductionID := "DB_OPTPLC_ExchangeData".PlcOptData.AUX_tPlatePacket.rgdProductionID[#TMP_dIndex];
           #INO_tCaps.tNewCapToInsert.rgtLites[#TMP_dIndex].strProdDescr := '';
           #INO_tCaps.tNewCapToInsert.rgtLites[#TMP_dIndex].dQualityID := "DB_OPTPLC_ExchangeData".PlcOptData.AUX_tPlatePacket.rgdQualityID[#TMP_dIndex];
           #INO_tCaps.tNewCapToInsert.rgtLites[#TMP_dIndex].strQualityDescr := '';
           #INO_tCaps.tNewCapToInsert.rgtLites[#TMP_dIndex].dCameraRecipeID := "DB_OPTPLC_ExchangeData".PlcOptData.AUX_tPlatePacket.dGeomID;
           #INO_tCaps.tNewCapToInsert.rgtLites[#TMP_dIndex].dWidth_cmm := "DB_OPTPLC_ExchangeData".PlcOptData.AUX_tPlatePacket.rgdLiteWidth_cmm[#TMP_dIndex];
           #INO_tCaps.tNewCapToInsert.rgtLites[#TMP_dIndex].dBarycentre_cmm := 0;
           #INO_tCaps.tNewCapToInsert.rgtLites[#TMP_dIndex].dCulletCause := "DB_OPTPLC_ExchangeData".PlcOptData.AUX_tPlatePacket.rgdCulletCause[#TMP_dIndex];
           #INO_tCaps.tNewCapToInsert.rgtLites[#TMP_dIndex].rgxLayers[0] := "DB_OPTPLC_ExchangeData".PlcOptData.AUX_tPlatePacket.rgtLiteFlags[#TMP_dIndex].xPow1Req;
           #INO_tCaps.tNewCapToInsert.rgtLites[#TMP_dIndex].rgxLayers[1] := "DB_OPTPLC_ExchangeData".PlcOptData.AUX_tPlatePacket.rgtLiteFlags[#TMP_dIndex].xPow2Req;
           #INO_tCaps.tNewCapToInsert.rgtLites[#TMP_dIndex].dMainDestination := "DB_OPTPLC_ExchangeData".PlcOptData.AUX_tPlatePacket.rgdDestMain[#TMP_dIndex];
           #INO_tCaps.tNewCapToInsert.rgtLites[#TMP_dIndex].dAltDestination := "DB_OPTPLC_ExchangeData".PlcOptData.AUX_tPlatePacket.rgdDestAlt[#TMP_dIndex];
           #INO_tCaps.tNewCapToInsert.rgtLites[#TMP_dIndex].d2ndDestionation := "DB_OPTPLC_ExchangeData".PlcOptData.AUX_tPlatePacket.rgdDest2Nd[#TMP_dIndex];

           #INO_tCaps.tNewCapToInsert.rgtLites[#TMP_dIndex].dMainDestination := "DB_OPTPLC_ExchangeData".PlcOptData.AUX_tPlatePacket.rgdDestMain[#TMP_dIndex];
           #INO_tCaps.tNewCapToInsert.rgtLites[#TMP_dIndex].dAltDestination := "DB_OPTPLC_ExchangeData".PlcOptData.AUX_tPlatePacket.rgdDestAlt[#TMP_dIndex];
           #INO_tCaps.tNewCapToInsert.rgtLites[#TMP_dIndex].d2ndDestionation := "DB_OPTPLC_ExchangeData".PlcOptData.AUX_tPlatePacket.rgdDest2Nd[#TMP_dIndex];

           #INO_tCaps.tNewCapToInsert.rgtLites[#TMP_dIndex].tRequests.dMapLaserHeadOp := 0;
           #INO_tCaps.tNewCapToInsert.rgtLites[#TMP_dIndex].tRequests.dMapLaserHeadOppOp := 0;
           #INO_tCaps.tNewCapToInsert.rgtLites[#TMP_dIndex].xSaturationPlate := "DB_OPTPLC_ExchangeData".PlcOptData.AUX_tPlatePacket.rgtLiteFlags[#TMP_dIndex].xSatPlate;
           #INO_tCaps.tNewCapToInsert.rgtLites[#TMP_dIndex].tRequests.xGeomInsp := "DB_OPTPLC_ExchangeData".PlcOptData.AUX_tPlatePacket.rgtLiteFlags[#TMP_dIndex].xGeomInsp;

       END_FOR;

       #INO_tCaps.xInsertCapOnTrack := TRUE;

   ELSIF "DB_OPTPLC_ExchangeData".PlcOptData.xCapDataReady THEN

       "DB_OPTPLC_ExchangeData".PlcOptData.xCapDataReady := FALSE;

   END_IF;
   *)
END_REGION

REGION Network 8 (SCL): Prepare the defects for internal plc optimizer
   (*
   IF "DB_OPTPLC_ExchangeData".TrackingData.tDefects.dNumOfDef = 0 AND #INO_tDefects.tDefectsforOptPlc.dNumberOfDefect > 0 THEN

       FOR #TMP_dIndex := 0 TO #INO_tDefects.tDefectsforOptPlc.dNumberOfDefect - 1 DO

           "DB_OPTPLC_ExchangeData".TrackingData.tDefects.rgtDefecList[#TMP_dIndex].dClass := #INO_tDefects.tDefectsforOptPlc.rgtDefects[#TMP_dIndex].dClass;
           "DB_OPTPLC_ExchangeData".TrackingData.tDefects.rgtDefecList[#TMP_dIndex].dSubtype := #INO_tDefects.tDefectsforOptPlc.rgtDefects[#TMP_dIndex].dSubType;
           "DB_OPTPLC_ExchangeData".TrackingData.tDefects.rgtDefecList[#TMP_dIndex].dPositionX_cmm := #INO_tDefects.tDefectsforOptPlc.rgtDefects[#TMP_dIndex].dXPosition_cmm;
           "DB_OPTPLC_ExchangeData".TrackingData.tDefects.rgtDefecList[#TMP_dIndex].dPositionY_cmm := #INO_tDefects.tDefectsforOptPlc.rgtDefects[#TMP_dIndex].dYPosition_cmm;
           "DB_OPTPLC_ExchangeData".TrackingData.tDefects.rgtDefecList[#TMP_dIndex].dLength_um := #INO_tDefects.tDefectsforOptPlc.rgtDefects[#TMP_dIndex].dTotalLength_um;
           "DB_OPTPLC_ExchangeData".TrackingData.tDefects.rgtDefecList[#TMP_dIndex].dWidth_um := #INO_tDefects.tDefectsforOptPlc.rgtDefects[#TMP_dIndex].dTotalWidth_um;

       END_FOR;

       "DB_OPTPLC_ExchangeData".TrackingData.tDefects.dNumOfDef := #INO_tDefects.tDefectsforOptPlc.dNumberOfDefect;
       #INO_tDefects.tDefectsforOptPlc.dNumberOfDefect := 0;

   END_IF;*)
END_REGION
END_FUNCTION_BLOCK

